(* Logix 5000 project; controller PLC_MCC1300_75F1 vendor 1 type 14 code 166 rev 32.11; software revision 32.04; part 15 of 83 *)
(* tags used below, declared in another part *)
   M302SpeedUp : MAC_SpeedUp;
   TMP_d : DINT;
   TMP_xPositioning : BOOL;
   TMP_xReverse : BOOL;
   TMP_xRun : BOOL;
   xAlwaysOFF : BOOL;
   Z300_Conveyor : UDT_StandConv[29];
   Z300_Conveyor_Conf : UDT_Conveyor_Config[29];
   Z300_Conveyor_HMW : MAC_Conveyor_ZC_HMW[29];
   Z300_Conveyor_IN_MOTION : MAC_Conveyor_ZC_IN_MOTION[29];
   Z301_HMR : MAC_Zone_ML_HMR;
(* CommandLogic, continued *)

ROUTINE M305M1_Conveyor_Output   (* ladder *)
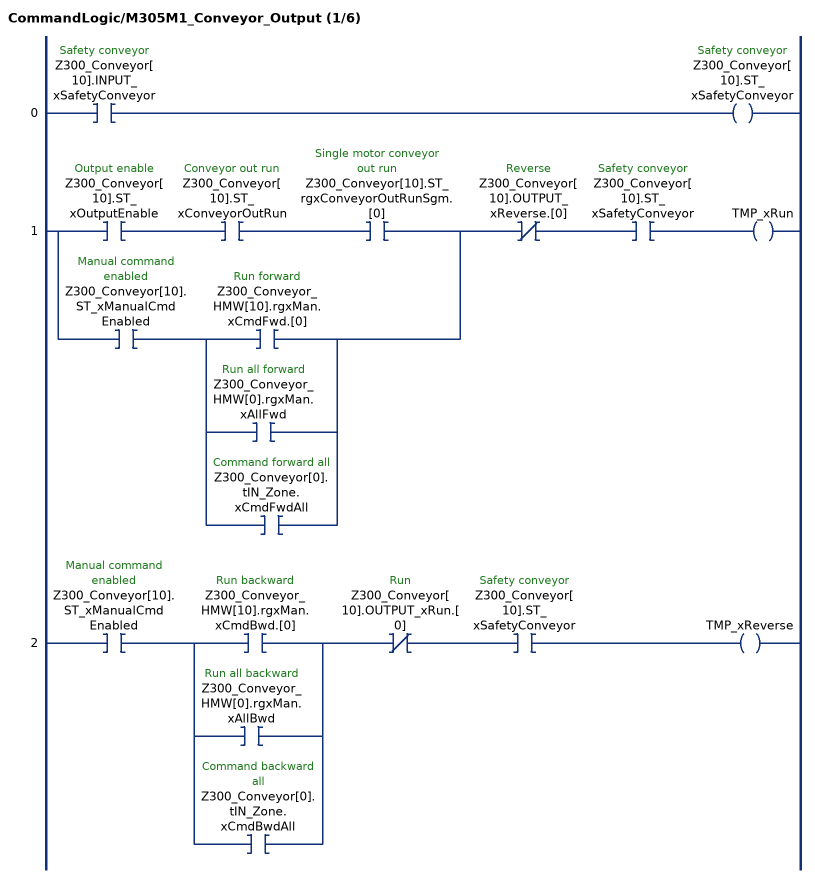
   0: XIC(Z300_Conveyor[10].INPUT_xSafetyConveyor)OTE(Z300_Conveyor[10].ST_xSafetyConveyor);
   1: [XIC(Z300_Conveyor[10].ST_xOutputEnable) XIC(Z300_Conveyor[10].ST_xConveyorOutRun) XIC(Z300_Conveyor[10].ST_rgxConveyorOutRunSgm.[0]) ,XIC(Z300_Conveyor[10].ST_xManualCmdEnabled) [XIC(Z300_Conveyor_HMW[10].rgxMan.xCmdFwd.[0]) ,XIC(Z300_Conveyor_HMW[0].rgxMan.xAllFwd) ,XIC(Z300_Conveyor[0].tIN_Zone.xCmdFwdAll) ] ]XIO(Z300_Conveyor[10].OUTPUT_xReverse.[0])XIC(Z300_Conveyor[10].ST_xSafetyConveyor)OTE(TMP_xRun);
   2: XIC(Z300_Conveyor[10].ST_xManualCmdEnabled)[XIC(Z300_Conveyor_HMW[10].rgxMan.xCmdBwd.[0]) ,XIC(Z300_Conveyor_HMW[0].rgxMan.xAllBwd) ,XIC(Z300_Conveyor[0].tIN_Zone.xCmdBwdAll) ]XIO(Z300_Conveyor[10].OUTPUT_xRun.[0])XIC(Z300_Conveyor[10].ST_xSafetyConveyor)OTE(TMP_xReverse);
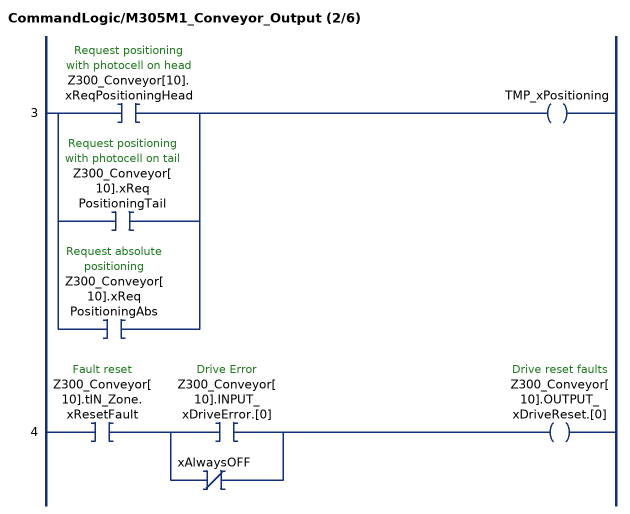
   3: [XIC(Z300_Conveyor[10].xReqPositioningHead) ,XIC(Z300_Conveyor[10].xReqPositioningTail) ,XIC(Z300_Conveyor[10].xReqPositioningAbs) ]OTE(TMP_xPositioning);
   4: XIC(Z300_Conveyor[10].tIN_Zone.xResetFault)[XIC(Z300_Conveyor[10].INPUT_xDriveError.[0]) ,XIO(xAlwaysOFF) ]OTE(Z300_Conveyor[10].OUTPUT_xDriveReset.[0]);
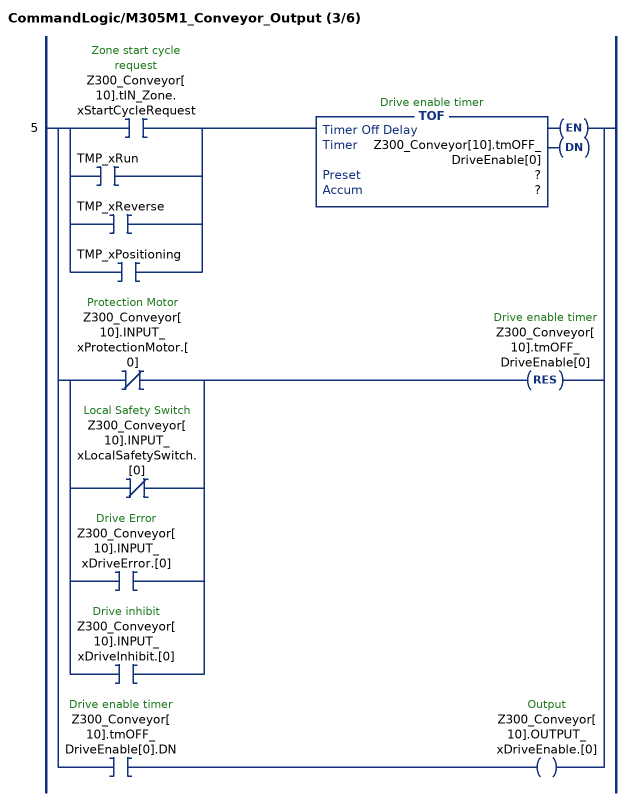
   5: [[XIC(Z300_Conveyor[10].tIN_Zone.xStartCycleRequest) ,XIC(TMP_xRun) ,XIC(TMP_xReverse) ,XIC(TMP_xPositioning) ] TOF(Z300_Conveyor[10].tmOFF_DriveEnable[0],?,?) ,[XIO(Z300_Conveyor[10].INPUT_xProtectionMotor.[0]) ,XIO(Z300_Conveyor[10].INPUT_xLocalSafetySwitch.[0]) ,XIC(Z300_Conveyor[10].INPUT_xDriveError.[0]) ,XIC(Z300_Conveyor[10].INPUT_xDriveInhibit.[0]) ] RES(Z300_Conveyor[10].tmOFF_DriveEnable[0]) ,XIC(Z300_Conveyor[10].tmOFF_DriveEnable[0].DN) OTE(Z300_Conveyor[10].OUTPUT_xDriveEnable.[0]) ];
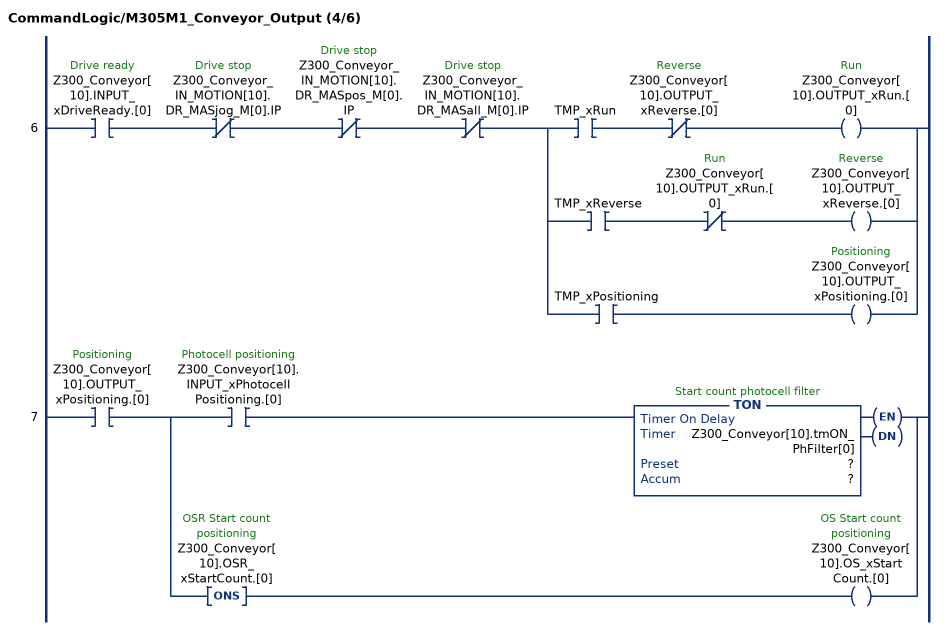
   6: XIC(Z300_Conveyor[10].INPUT_xDriveReady.[0])XIO(Z300_Conveyor_IN_MOTION[10].DR_MASjog_M[0].IP)XIO(Z300_Conveyor_IN_MOTION[10].DR_MASpos_M[0].IP)XIO(Z300_Conveyor_IN_MOTION[10].DR_MASall_M[0].IP)[XIC(TMP_xRun) XIO(Z300_Conveyor[10].OUTPUT_xReverse.[0]) OTE(Z300_Conveyor[10].OUTPUT_xRun.[0]) ,XIC(TMP_xReverse) XIO(Z300_Conveyor[10].OUTPUT_xRun.[0]) OTE(Z300_Conveyor[10].OUTPUT_xReverse.[0]) ,XIC(TMP_xPositioning) OTE(Z300_Conveyor[10].OUTPUT_xPositioning.[0]) ];
   7: XIC(Z300_Conveyor[10].OUTPUT_xPositioning.[0])[XIC(Z300_Conveyor[10].INPUT_xPhotocellPositioning.[0]) TON(Z300_Conveyor[10].tmON_PhFilter[0],?,?) ,ONS(Z300_Conveyor[10].OSR_xStartCount.[0]) OTE(Z300_Conveyor[10].OS_xStartCount.[0]) ];
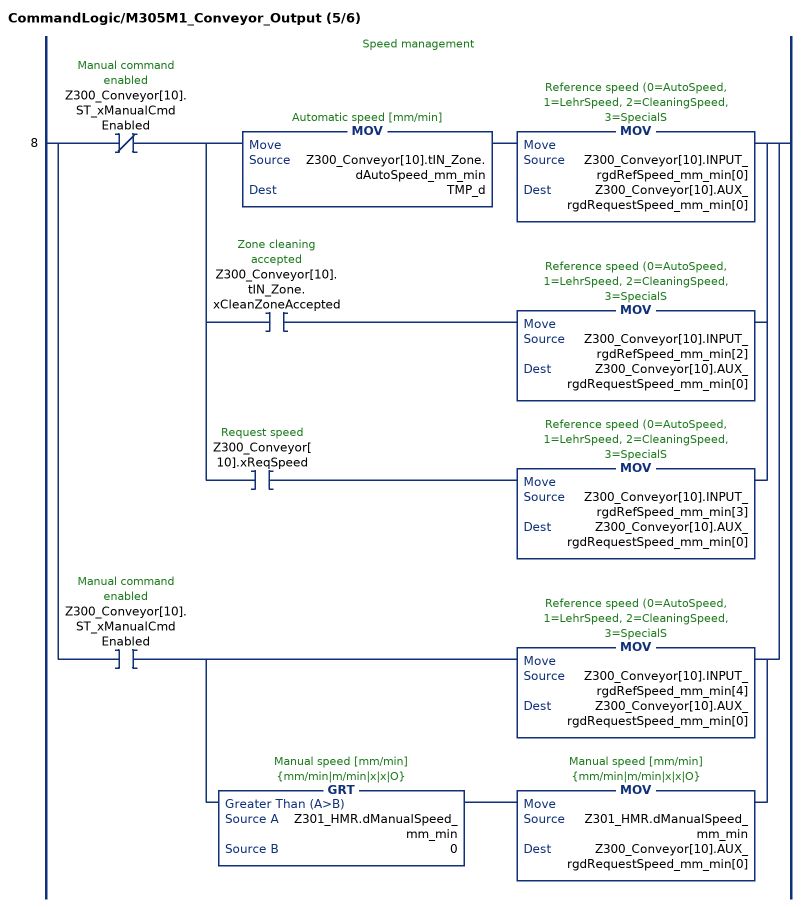
   // Speed management
   8: [XIO(Z300_Conveyor[10].ST_xManualCmdEnabled) [MOV(Z300_Conveyor[10].tIN_Zone.dAutoSpeed_mm_min,TMP_d) MOV(Z300_Conveyor[10].INPUT_rgdRefSpeed_mm_min[0],Z300_Conveyor[10].AUX_rgdRequestSpeed_mm_min[0]) ,XIC(Z300_Conveyor[10].tIN_Zone.xCleanZoneAccepted) MOV(Z300_Conveyor[10].INPUT_rgdRefSpeed_mm_min[2],Z300_Conveyor[10].AUX_rgdRequestSpeed_mm_min[0]) ,XIC(Z300_Conveyor[10].xReqSpeed) MOV(Z300_Conveyor[10].INPUT_rgdRefSpeed_mm_min[3],Z300_Conveyor[10].AUX_rgdRequestSpeed_mm_min[0]) ] ,XIC(Z300_Conveyor[10].ST_xManualCmdEnabled) [MOV(Z300_Conveyor[10].INPUT_rgdRefSpeed_mm_min[4],Z300_Conveyor[10].AUX_rgdRequestSpeed_mm_min[0]) ,GRT(Z301_HMR.dManualSpeed_mm_min,0) MOV(Z301_HMR.dManualSpeed_mm_min,Z300_Conveyor[10].AUX_rgdRequestSpeed_mm_min[0]) ] ];
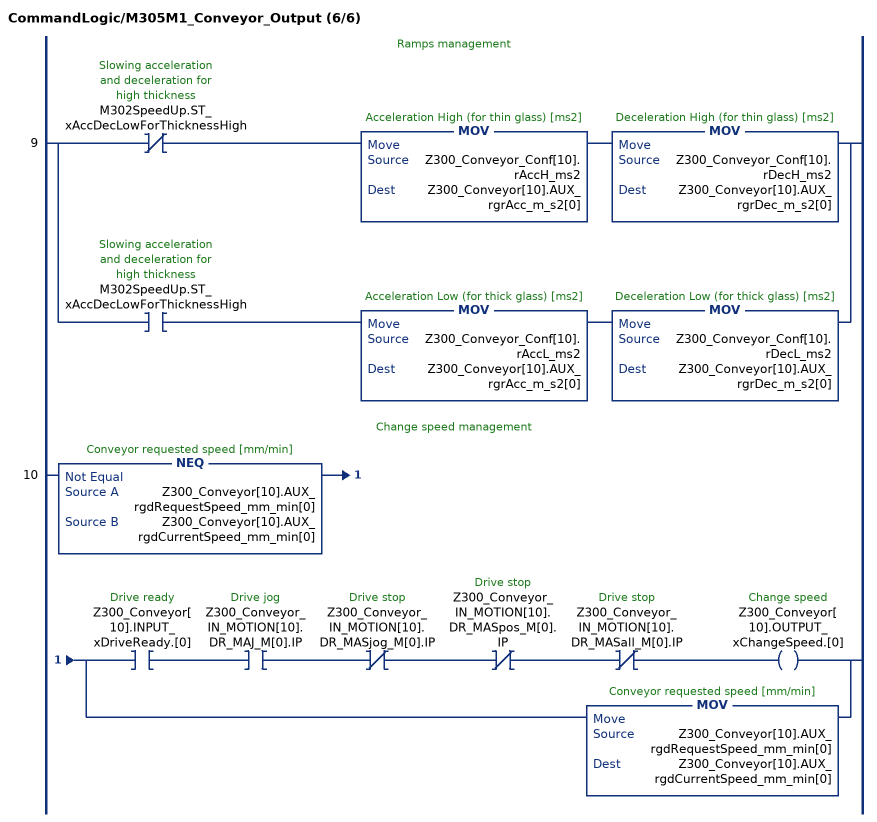
   // Ramps management
   9: [XIO(M302SpeedUp.ST_xAccDecLowForThicknessHigh) MOV(Z300_Conveyor_Conf[10].rAccH_ms2,Z300_Conveyor[10].AUX_rgrAcc_m_s2[0]) MOV(Z300_Conveyor_Conf[10].rDecH_ms2,Z300_Conveyor[10].AUX_rgrDec_m_s2[0]) ,XIC(M302SpeedUp.ST_xAccDecLowForThicknessHigh) MOV(Z300_Conveyor_Conf[10].rAccL_ms2,Z300_Conveyor[10].AUX_rgrAcc_m_s2[0]) MOV(Z300_Conveyor_Conf[10].rDecL_ms2,Z300_Conveyor[10].AUX_rgrDec_m_s2[0]) ];
   // Change speed management
   10: NEQ(Z300_Conveyor[10].AUX_rgdRequestSpeed_mm_min[0],Z300_Conveyor[10].AUX_rgdCurrentSpeed_mm_min[0])[XIC(Z300_Conveyor[10].INPUT_xDriveReady.[0]) XIC(Z300_Conveyor_IN_MOTION[10].DR_MAJ_M[0].IP) XIO(Z300_Conveyor_IN_MOTION[10].DR_MASjog_M[0].IP) XIO(Z300_Conveyor_IN_MOTION[10].DR_MASpos_M[0].IP) XIO(Z300_Conveyor_IN_MOTION[10].DR_MASall_M[0].IP) OTE(Z300_Conveyor[10].OUTPUT_xChangeSpeed.[0]) ,MOV(Z300_Conveyor[10].AUX_rgdRequestSpeed_mm_min[0],Z300_Conveyor[10].AUX_rgdCurrentSpeed_mm_min[0]) ];
END_ROUTINE

ROUTINE M306M1_Conveyor_Output   (* ladder *)
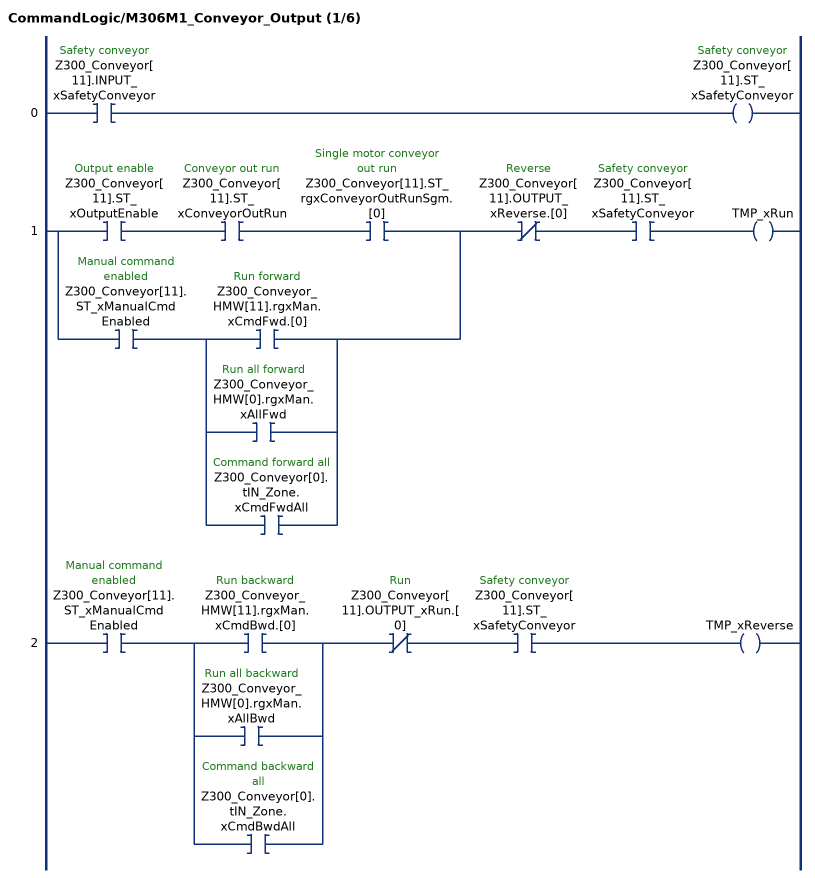
   0: XIC(Z300_Conveyor[11].INPUT_xSafetyConveyor)OTE(Z300_Conveyor[11].ST_xSafetyConveyor);
   1: [XIC(Z300_Conveyor[11].ST_xOutputEnable) XIC(Z300_Conveyor[11].ST_xConveyorOutRun) XIC(Z300_Conveyor[11].ST_rgxConveyorOutRunSgm.[0]) ,XIC(Z300_Conveyor[11].ST_xManualCmdEnabled) [XIC(Z300_Conveyor_HMW[11].rgxMan.xCmdFwd.[0]) ,XIC(Z300_Conveyor_HMW[0].rgxMan.xAllFwd) ,XIC(Z300_Conveyor[0].tIN_Zone.xCmdFwdAll) ] ]XIO(Z300_Conveyor[11].OUTPUT_xReverse.[0])XIC(Z300_Conveyor[11].ST_xSafetyConveyor)OTE(TMP_xRun);
   2: XIC(Z300_Conveyor[11].ST_xManualCmdEnabled)[XIC(Z300_Conveyor_HMW[11].rgxMan.xCmdBwd.[0]) ,XIC(Z300_Conveyor_HMW[0].rgxMan.xAllBwd) ,XIC(Z300_Conveyor[0].tIN_Zone.xCmdBwdAll) ]XIO(Z300_Conveyor[11].OUTPUT_xRun.[0])XIC(Z300_Conveyor[11].ST_xSafetyConveyor)OTE(TMP_xReverse);
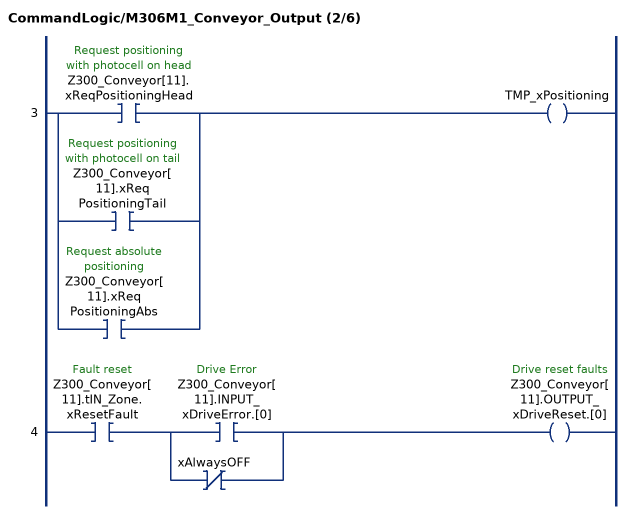
   3: [XIC(Z300_Conveyor[11].xReqPositioningHead) ,XIC(Z300_Conveyor[11].xReqPositioningTail) ,XIC(Z300_Conveyor[11].xReqPositioningAbs) ]OTE(TMP_xPositioning);
   4: XIC(Z300_Conveyor[11].tIN_Zone.xResetFault)[XIC(Z300_Conveyor[11].INPUT_xDriveError.[0]) ,XIO(xAlwaysOFF) ]OTE(Z300_Conveyor[11].OUTPUT_xDriveReset.[0]);
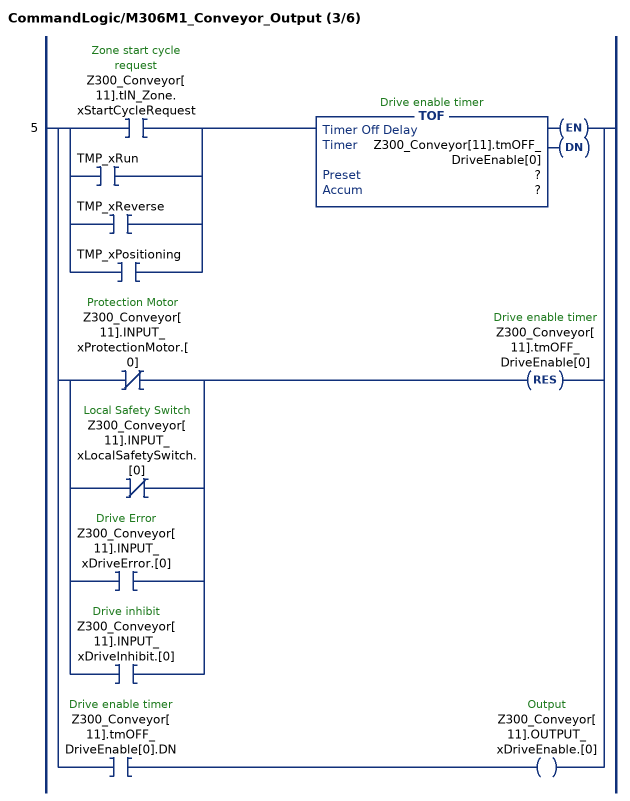
   5: [[XIC(Z300_Conveyor[11].tIN_Zone.xStartCycleRequest) ,XIC(TMP_xRun) ,XIC(TMP_xReverse) ,XIC(TMP_xPositioning) ] TOF(Z300_Conveyor[11].tmOFF_DriveEnable[0],?,?) ,[XIO(Z300_Conveyor[11].INPUT_xProtectionMotor.[0]) ,XIO(Z300_Conveyor[11].INPUT_xLocalSafetySwitch.[0]) ,XIC(Z300_Conveyor[11].INPUT_xDriveError.[0]) ,XIC(Z300_Conveyor[11].INPUT_xDriveInhibit.[0]) ] RES(Z300_Conveyor[11].tmOFF_DriveEnable[0]) ,XIC(Z300_Conveyor[11].tmOFF_DriveEnable[0].DN) OTE(Z300_Conveyor[11].OUTPUT_xDriveEnable.[0]) ];
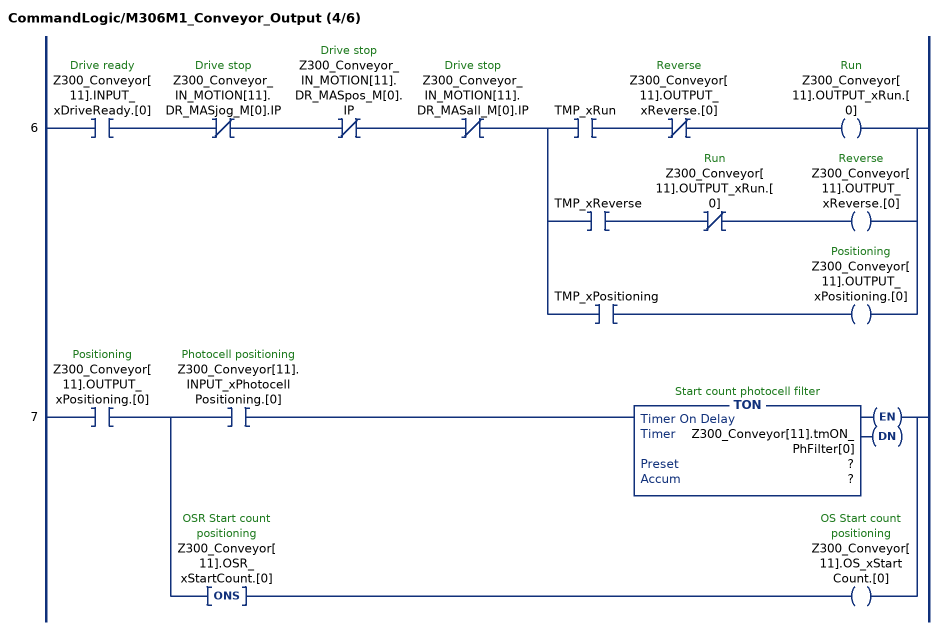
   6: XIC(Z300_Conveyor[11].INPUT_xDriveReady.[0])XIO(Z300_Conveyor_IN_MOTION[11].DR_MASjog_M[0].IP)XIO(Z300_Conveyor_IN_MOTION[11].DR_MASpos_M[0].IP)XIO(Z300_Conveyor_IN_MOTION[11].DR_MASall_M[0].IP)[XIC(TMP_xRun) XIO(Z300_Conveyor[11].OUTPUT_xReverse.[0]) OTE(Z300_Conveyor[11].OUTPUT_xRun.[0]) ,XIC(TMP_xReverse) XIO(Z300_Conveyor[11].OUTPUT_xRun.[0]) OTE(Z300_Conveyor[11].OUTPUT_xReverse.[0]) ,XIC(TMP_xPositioning) OTE(Z300_Conveyor[11].OUTPUT_xPositioning.[0]) ];
   7: XIC(Z300_Conveyor[11].OUTPUT_xPositioning.[0])[XIC(Z300_Conveyor[11].INPUT_xPhotocellPositioning.[0]) TON(Z300_Conveyor[11].tmON_PhFilter[0],?,?) ,ONS(Z300_Conveyor[11].OSR_xStartCount.[0]) OTE(Z300_Conveyor[11].OS_xStartCount.[0]) ];
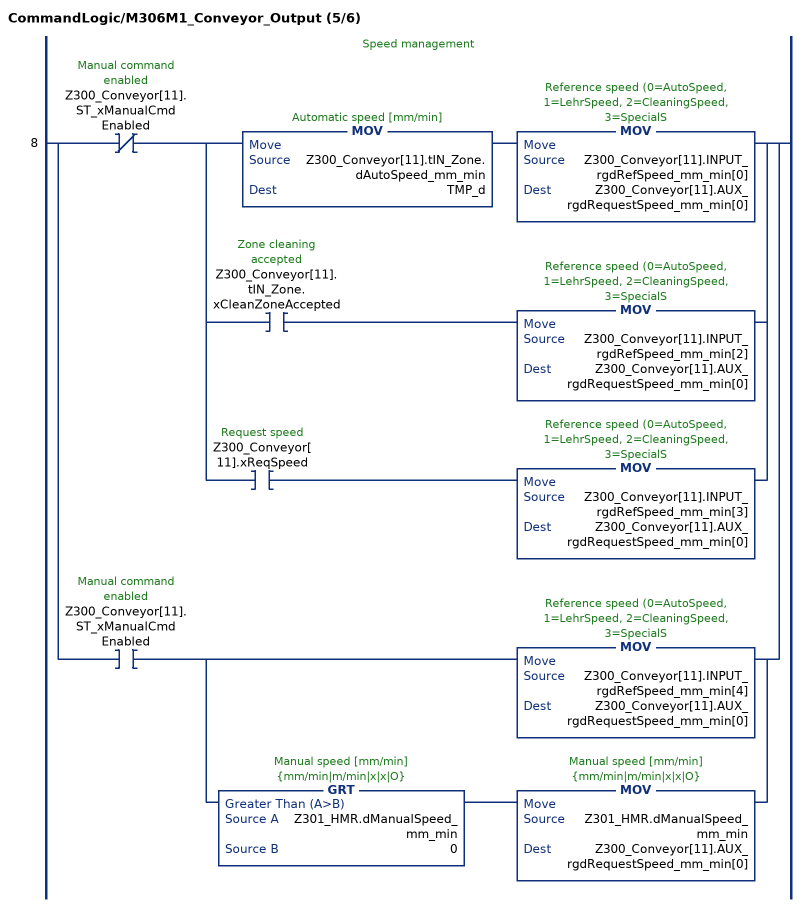
   // Speed management
   8: [XIO(Z300_Conveyor[11].ST_xManualCmdEnabled) [MOV(Z300_Conveyor[11].tIN_Zone.dAutoSpeed_mm_min,TMP_d) MOV(Z300_Conveyor[11].INPUT_rgdRefSpeed_mm_min[0],Z300_Conveyor[11].AUX_rgdRequestSpeed_mm_min[0]) ,XIC(Z300_Conveyor[11].tIN_Zone.xCleanZoneAccepted) MOV(Z300_Conveyor[11].INPUT_rgdRefSpeed_mm_min[2],Z300_Conveyor[11].AUX_rgdRequestSpeed_mm_min[0]) ,XIC(Z300_Conveyor[11].xReqSpeed) MOV(Z300_Conveyor[11].INPUT_rgdRefSpeed_mm_min[3],Z300_Conveyor[11].AUX_rgdRequestSpeed_mm_min[0]) ] ,XIC(Z300_Conveyor[11].ST_xManualCmdEnabled) [MOV(Z300_Conveyor[11].INPUT_rgdRefSpeed_mm_min[4],Z300_Conveyor[11].AUX_rgdRequestSpeed_mm_min[0]) ,GRT(Z301_HMR.dManualSpeed_mm_min,0) MOV(Z301_HMR.dManualSpeed_mm_min,Z300_Conveyor[11].AUX_rgdRequestSpeed_mm_min[0]) ] ];
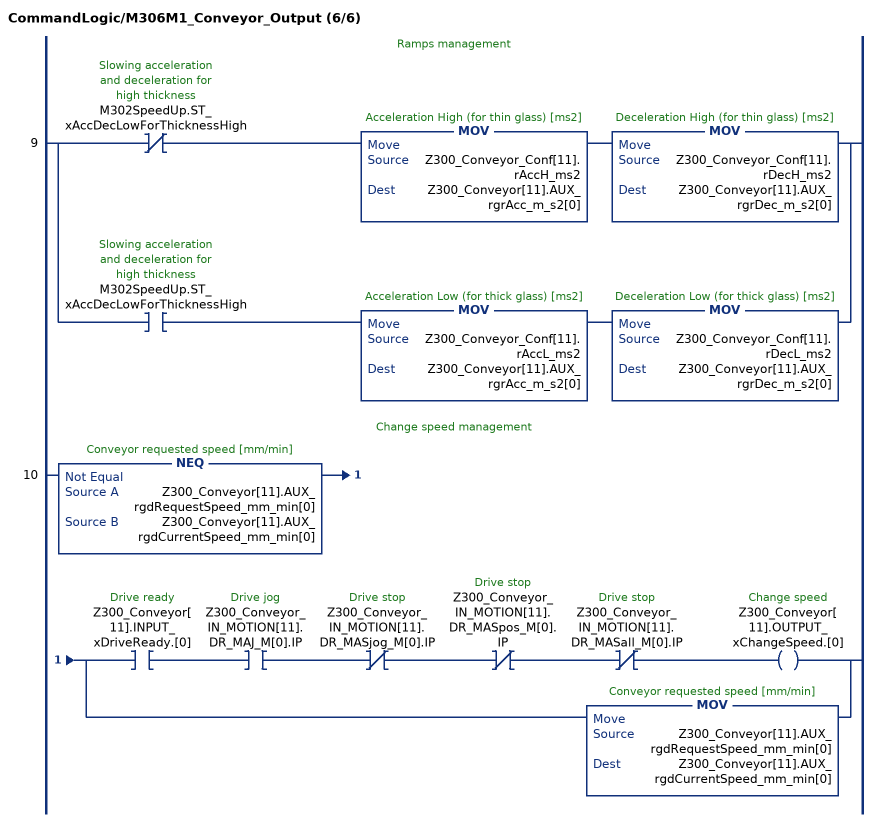
   // Ramps management
   9: [XIO(M302SpeedUp.ST_xAccDecLowForThicknessHigh) MOV(Z300_Conveyor_Conf[11].rAccH_ms2,Z300_Conveyor[11].AUX_rgrAcc_m_s2[0]) MOV(Z300_Conveyor_Conf[11].rDecH_ms2,Z300_Conveyor[11].AUX_rgrDec_m_s2[0]) ,XIC(M302SpeedUp.ST_xAccDecLowForThicknessHigh) MOV(Z300_Conveyor_Conf[11].rAccL_ms2,Z300_Conveyor[11].AUX_rgrAcc_m_s2[0]) MOV(Z300_Conveyor_Conf[11].rDecL_ms2,Z300_Conveyor[11].AUX_rgrDec_m_s2[0]) ];
   // Change speed management
   10: NEQ(Z300_Conveyor[11].AUX_rgdRequestSpeed_mm_min[0],Z300_Conveyor[11].AUX_rgdCurrentSpeed_mm_min[0])[XIC(Z300_Conveyor[11].INPUT_xDriveReady.[0]) XIC(Z300_Conveyor_IN_MOTION[11].DR_MAJ_M[0].IP) XIO(Z300_Conveyor_IN_MOTION[11].DR_MASjog_M[0].IP) XIO(Z300_Conveyor_IN_MOTION[11].DR_MASpos_M[0].IP) XIO(Z300_Conveyor_IN_MOTION[11].DR_MASall_M[0].IP) OTE(Z300_Conveyor[11].OUTPUT_xChangeSpeed.[0]) ,MOV(Z300_Conveyor[11].AUX_rgdRequestSpeed_mm_min[0],Z300_Conveyor[11].AUX_rgdCurrentSpeed_mm_min[0]) ];
END_ROUTINE

ROUTINE M307AM1_Conveyor_Output   (* ladder *)
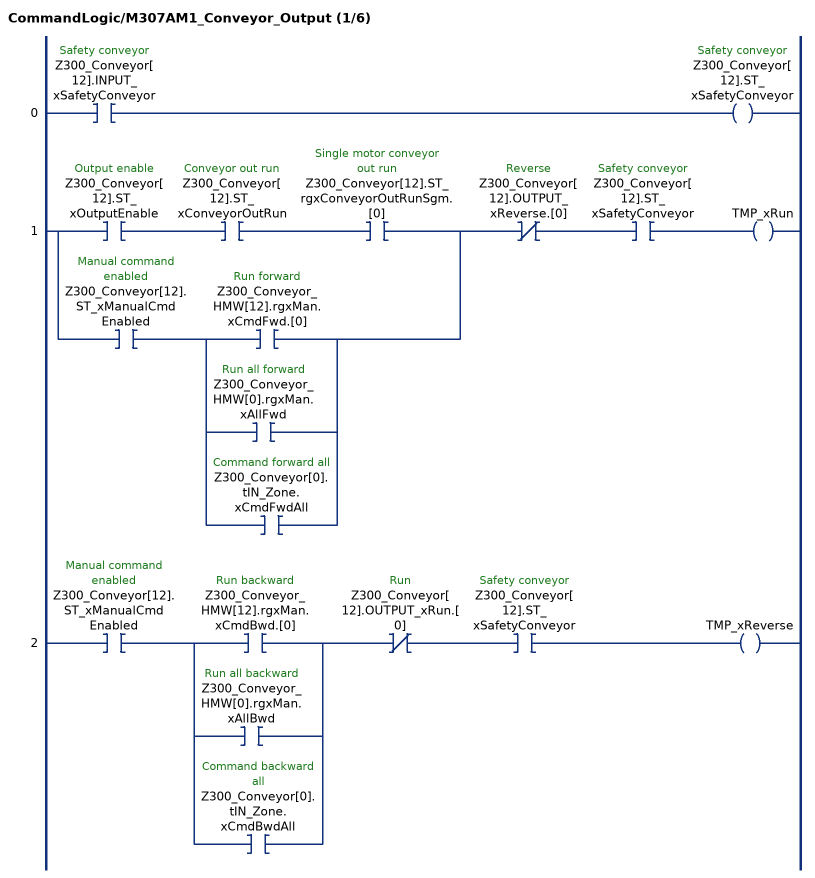
   0: XIC(Z300_Conveyor[12].INPUT_xSafetyConveyor)OTE(Z300_Conveyor[12].ST_xSafetyConveyor);
   1: [XIC(Z300_Conveyor[12].ST_xOutputEnable) XIC(Z300_Conveyor[12].ST_xConveyorOutRun) XIC(Z300_Conveyor[12].ST_rgxConveyorOutRunSgm.[0]) ,XIC(Z300_Conveyor[12].ST_xManualCmdEnabled) [XIC(Z300_Conveyor_HMW[12].rgxMan.xCmdFwd.[0]) ,XIC(Z300_Conveyor_HMW[0].rgxMan.xAllFwd) ,XIC(Z300_Conveyor[0].tIN_Zone.xCmdFwdAll) ] ]XIO(Z300_Conveyor[12].OUTPUT_xReverse.[0])XIC(Z300_Conveyor[12].ST_xSafetyConveyor)OTE(TMP_xRun);
   2: XIC(Z300_Conveyor[12].ST_xManualCmdEnabled)[XIC(Z300_Conveyor_HMW[12].rgxMan.xCmdBwd.[0]) ,XIC(Z300_Conveyor_HMW[0].rgxMan.xAllBwd) ,XIC(Z300_Conveyor[0].tIN_Zone.xCmdBwdAll) ]XIO(Z300_Conveyor[12].OUTPUT_xRun.[0])XIC(Z300_Conveyor[12].ST_xSafetyConveyor)OTE(TMP_xReverse);
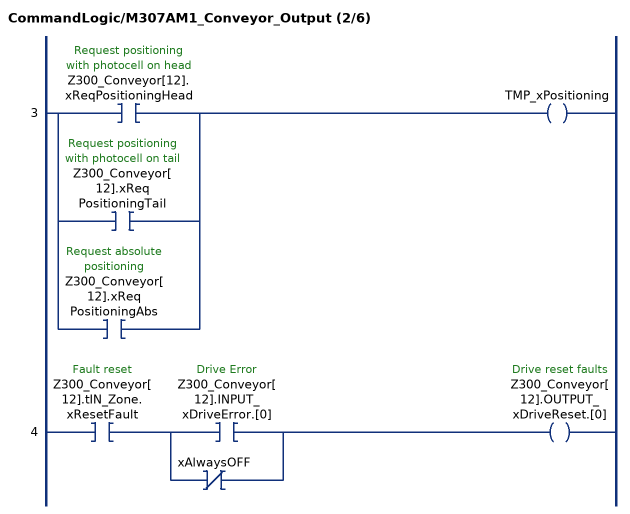
   3: [XIC(Z300_Conveyor[12].xReqPositioningHead) ,XIC(Z300_Conveyor[12].xReqPositioningTail) ,XIC(Z300_Conveyor[12].xReqPositioningAbs) ]OTE(TMP_xPositioning);
   4: XIC(Z300_Conveyor[12].tIN_Zone.xResetFault)[XIC(Z300_Conveyor[12].INPUT_xDriveError.[0]) ,XIO(xAlwaysOFF) ]OTE(Z300_Conveyor[12].OUTPUT_xDriveReset.[0]);
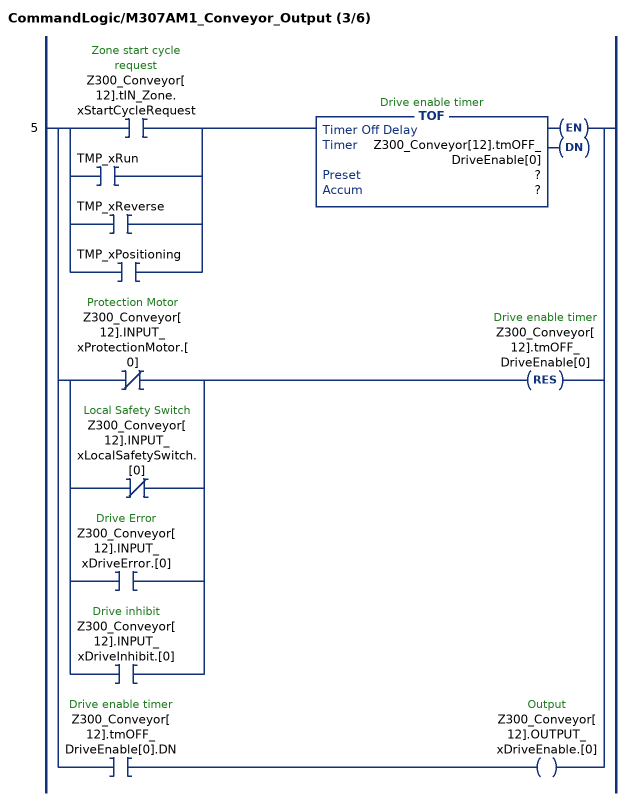
   5: [[XIC(Z300_Conveyor[12].tIN_Zone.xStartCycleRequest) ,XIC(TMP_xRun) ,XIC(TMP_xReverse) ,XIC(TMP_xPositioning) ] TOF(Z300_Conveyor[12].tmOFF_DriveEnable[0],?,?) ,[XIO(Z300_Conveyor[12].INPUT_xProtectionMotor.[0]) ,XIO(Z300_Conveyor[12].INPUT_xLocalSafetySwitch.[0]) ,XIC(Z300_Conveyor[12].INPUT_xDriveError.[0]) ,XIC(Z300_Conveyor[12].INPUT_xDriveInhibit.[0]) ] RES(Z300_Conveyor[12].tmOFF_DriveEnable[0]) ,XIC(Z300_Conveyor[12].tmOFF_DriveEnable[0].DN) OTE(Z300_Conveyor[12].OUTPUT_xDriveEnable.[0]) ];
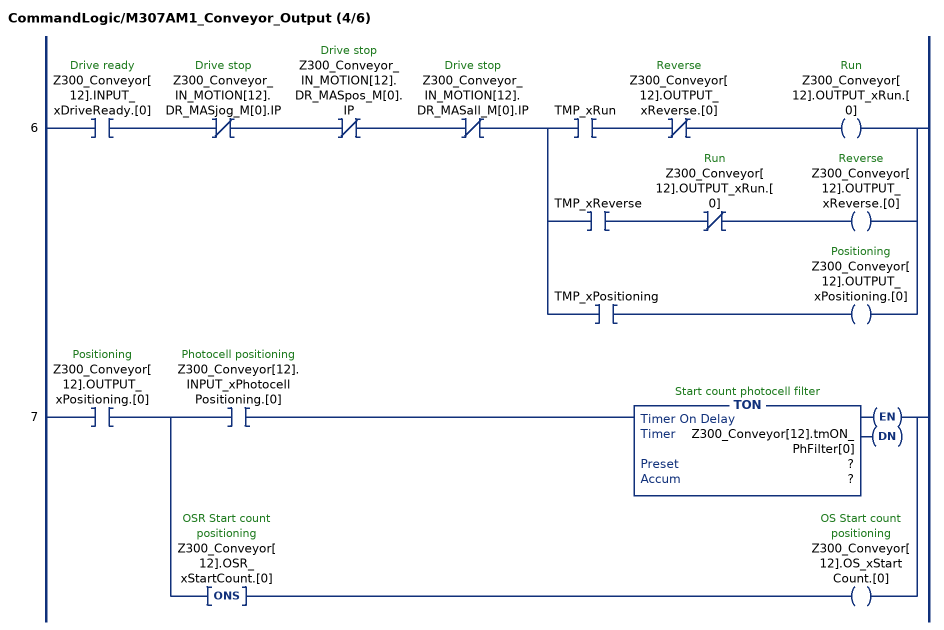
   6: XIC(Z300_Conveyor[12].INPUT_xDriveReady.[0])XIO(Z300_Conveyor_IN_MOTION[12].DR_MASjog_M[0].IP)XIO(Z300_Conveyor_IN_MOTION[12].DR_MASpos_M[0].IP)XIO(Z300_Conveyor_IN_MOTION[12].DR_MASall_M[0].IP)[XIC(TMP_xRun) XIO(Z300_Conveyor[12].OUTPUT_xReverse.[0]) OTE(Z300_Conveyor[12].OUTPUT_xRun.[0]) ,XIC(TMP_xReverse) XIO(Z300_Conveyor[12].OUTPUT_xRun.[0]) OTE(Z300_Conveyor[12].OUTPUT_xReverse.[0]) ,XIC(TMP_xPositioning) OTE(Z300_Conveyor[12].OUTPUT_xPositioning.[0]) ];
   7: XIC(Z300_Conveyor[12].OUTPUT_xPositioning.[0])[XIC(Z300_Conveyor[12].INPUT_xPhotocellPositioning.[0]) TON(Z300_Conveyor[12].tmON_PhFilter[0],?,?) ,ONS(Z300_Conveyor[12].OSR_xStartCount.[0]) OTE(Z300_Conveyor[12].OS_xStartCount.[0]) ];
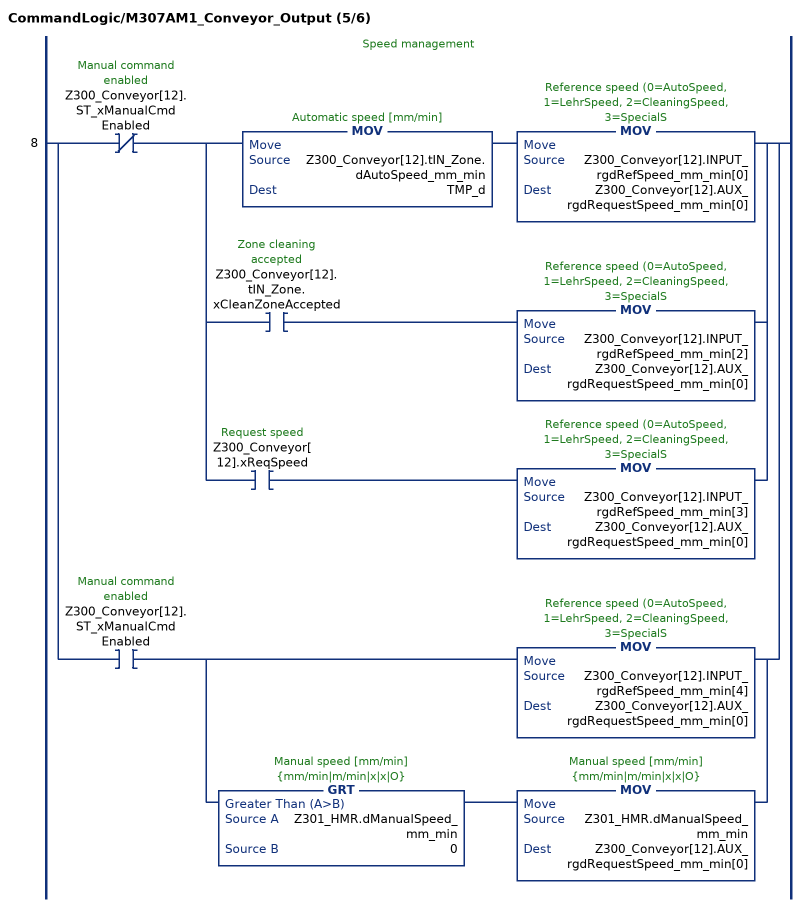
   // Speed management
   8: [XIO(Z300_Conveyor[12].ST_xManualCmdEnabled) [MOV(Z300_Conveyor[12].tIN_Zone.dAutoSpeed_mm_min,TMP_d) MOV(Z300_Conveyor[12].INPUT_rgdRefSpeed_mm_min[0],Z300_Conveyor[12].AUX_rgdRequestSpeed_mm_min[0]) ,XIC(Z300_Conveyor[12].tIN_Zone.xCleanZoneAccepted) MOV(Z300_Conveyor[12].INPUT_rgdRefSpeed_mm_min[2],Z300_Conveyor[12].AUX_rgdRequestSpeed_mm_min[0]) ,XIC(Z300_Conveyor[12].xReqSpeed) MOV(Z300_Conveyor[12].INPUT_rgdRefSpeed_mm_min[3],Z300_Conveyor[12].AUX_rgdRequestSpeed_mm_min[0]) ] ,XIC(Z300_Conveyor[12].ST_xManualCmdEnabled) [MOV(Z300_Conveyor[12].INPUT_rgdRefSpeed_mm_min[4],Z300_Conveyor[12].AUX_rgdRequestSpeed_mm_min[0]) ,GRT(Z301_HMR.dManualSpeed_mm_min,0) MOV(Z301_HMR.dManualSpeed_mm_min,Z300_Conveyor[12].AUX_rgdRequestSpeed_mm_min[0]) ] ];
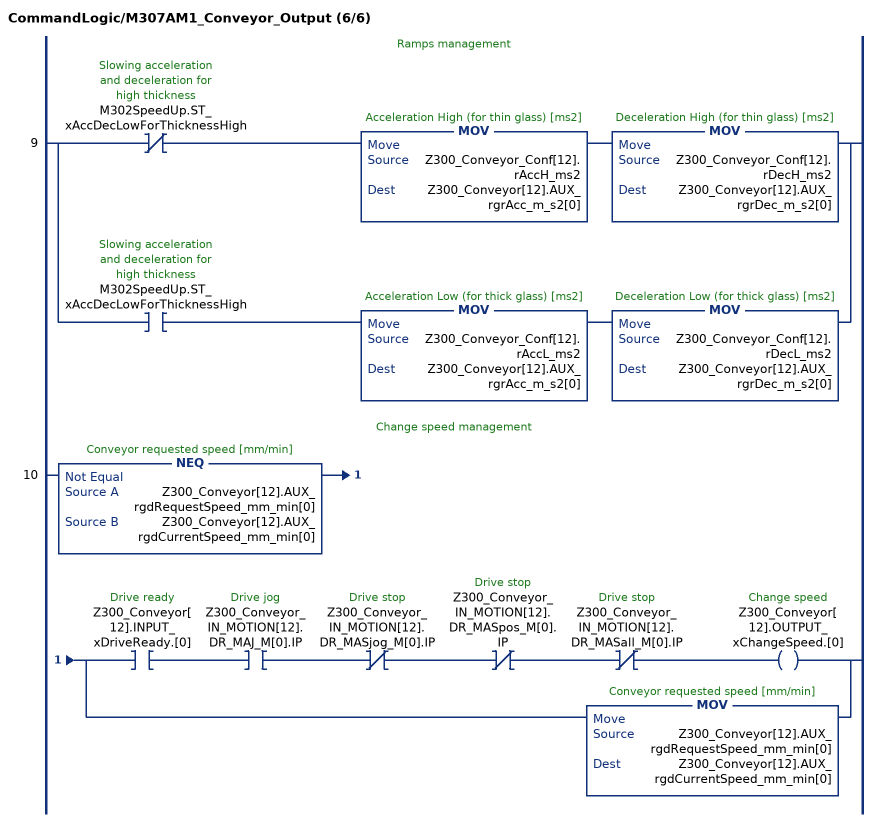
   // Ramps management
   9: [XIO(M302SpeedUp.ST_xAccDecLowForThicknessHigh) MOV(Z300_Conveyor_Conf[12].rAccH_ms2,Z300_Conveyor[12].AUX_rgrAcc_m_s2[0]) MOV(Z300_Conveyor_Conf[12].rDecH_ms2,Z300_Conveyor[12].AUX_rgrDec_m_s2[0]) ,XIC(M302SpeedUp.ST_xAccDecLowForThicknessHigh) MOV(Z300_Conveyor_Conf[12].rAccL_ms2,Z300_Conveyor[12].AUX_rgrAcc_m_s2[0]) MOV(Z300_Conveyor_Conf[12].rDecL_ms2,Z300_Conveyor[12].AUX_rgrDec_m_s2[0]) ];
   // Change speed management
   10: NEQ(Z300_Conveyor[12].AUX_rgdRequestSpeed_mm_min[0],Z300_Conveyor[12].AUX_rgdCurrentSpeed_mm_min[0])[XIC(Z300_Conveyor[12].INPUT_xDriveReady.[0]) XIC(Z300_Conveyor_IN_MOTION[12].DR_MAJ_M[0].IP) XIO(Z300_Conveyor_IN_MOTION[12].DR_MASjog_M[0].IP) XIO(Z300_Conveyor_IN_MOTION[12].DR_MASpos_M[0].IP) XIO(Z300_Conveyor_IN_MOTION[12].DR_MASall_M[0].IP) OTE(Z300_Conveyor[12].OUTPUT_xChangeSpeed.[0]) ,MOV(Z300_Conveyor[12].AUX_rgdRequestSpeed_mm_min[0],Z300_Conveyor[12].AUX_rgdCurrentSpeed_mm_min[0]) ];
END_ROUTINE
